   "Carrier_49_Slot2_Input" AT %IW2814 : Word;   // SLOT 2 INPUT WORD
   "Carrier_49_CrashDetectSW" AT %I2814.0 : Bool;   // CRASH DETECT SW
   "Carrier_49_SpareSafetyInput(2_1)" AT %I2814.1 : Bool;   // SPARE SAFETY INPUT
   "Carrier_49_SpareSafetyInput(2_2)" AT %I2814.2 : Bool;   // SPARE SAFETY INPUT
   "Carrier_49_SpareSafetyInput(2_3)" AT %I2814.3 : Bool;   // SPARE SAFETY INPUT
   "Carrier_49_SpareSafetyInput(2_4)" AT %I2814.4 : Bool;   // SPARE SAFETY INPUT
   "Carrier_49_SpareSafetyInput(2_5)" AT %I2814.5 : Bool;   // SPARE SAFETY INPUT
   "Carrier_49_SpareSafetyInput(2_6)" AT %I2814.6 : Bool;   // SPARE SAFETY INPUT
   "Carrier_49_SpareSafetyInput(2_7)" AT %I2814.7 : Bool;   // SPARE SAFETY INPUT
   "Carrier_49_Slot3_SafetyOutput" AT %IW2815 : Word;   // SLOT 3 SAFETY OUTPUT WORD
   "Carrier_49_Crash_Detect_OK" AT %I2815.0 : Bool;   // CARRIER CRASH DETECT
   "Carrier_49_SpareSafetyOutput(3_1)" AT %I2815.1 : Bool;   // SPARE SAFETY OUTPUT
   "Carrier_49_SpareSafetyOutput(3_2)" AT %I2815.2 : Bool;   // SPARE SAFETY OUTPUT
   "Carrier_49_SpareSafetyOutput(3_3)" AT %I2815.3 : Bool;   // SPARE SAFETY OUTPUT
   "Carrier_49_SpareSafetyOutput(3_4)" AT %I2815.4 : Bool;   // SPARE SAFETY OUTPUT
   "Carrier_49_SpareSafetyOutput(3_5)" AT %I2815.5 : Bool;   // SPARE SAFETY OUTPUT
   "Carrier_49_SpareSafetyOutput(3_6)" AT %I2815.6 : Bool;   // SPARE SAFETY OUTPUT
   "Carrier_49_SpareSafetyOutput(3_7)" AT %I2815.7 : Bool;   // SPARE SAFETY OUTPUT
   "Carrier_49_Slot4_Input" AT %IW2816 : Word;   // SLOT 4 INPUT WORD
   "Carrier_49_480VPowerOn_MDCB1" AT %I2816.0 : Bool;   // 480 VAC POWER ON MDCB 1
   "Carrier_49_SpareInput(4_1)" AT %I2816.1 : Bool;   // SPARE INPUT
   "Carrier_49_SpareInput(4_2)" AT %I2816.2 : Bool;   // SPARE INPUT
   "Carrier_49_SitopSelectStatus" AT %I2816.3 : Bool;   // SITOP SELECT STATUS
   "Carrier_49_DCsupplyOnPSCB2" AT %I2816.4 : Bool;   // DC SUPPLY ON PSCB 2
   "Carrier_49_SpareInput(4_5)" AT %I2816.5 : Bool;   // SPARE INPUT
   "Carrier_49_SpareInput(4_6)" AT %I2816.6 : Bool;   // SPARE INPUT
   "Carrier_49_SpareInput(4_7)" AT %I2816.7 : Bool;   // SPARE INPUT
   "Carrier_49_PB1_ProdHoldLH" AT %I2817.0 : Bool;   // PB 1 PRODUCTION HOLD LH
   "Carrier_49_PB2_ResetLH" AT %I2817.1 : Bool;   // PB 2 RESET LH
   "Carrier_49_PB3_ProdHoldRH" AT %I2817.2 : Bool;   // PB 3 PRODUCTION HOLD RH
   "Carrier_49_PB4_ResetRH" AT %I2817.3 : Bool;   // PB 4 RESET RH
   "Carrier_49_SpareInput(4_14)" AT %I2817.4 : Bool;   // SPARE INPUT
   "Carrier_49_SpareInput(4_15)" AT %I2817.5 : Bool;   // SPARE INPUT
   "Carrier_49_SpareInput(4_16)" AT %I2817.6 : Bool;   // SPARE INPUT
   "Carrier_49_SpareInput(4_17)" AT %I2817.7 : Bool;   // SPARE INPUT
   "Carrier_49_Slot5_Output" AT %IW2818 : Word;   // SLOT 5 OUTPUT WORD
   "Carrier_49_IRD400_HMI_24VDC_ENABLE" AT %I2818.0 : Bool;   // IRD 400 PANEL HMI 24V DC POWER
   "Carrier_49_FaultLight_LH" AT %I2818.1 : Bool;   // FAULT LIGHT LH
   "Carrier_49_RunLight_LH" AT %I2818.2 : Bool;   // RUN LIGHT LH
   "Carrier_49_FaultLight_RH" AT %I2818.3 : Bool;   // FAULT LIGHT RH
   "Carrier_49_RunLight_RH" AT %I2818.4 : Bool;   // RUN LIGHT RH
   "Carrier_49_SpareOutput(5_5)" AT %I2818.5 : Bool;   // SPARE OUTPUT
   "Carrier_49_SpareOutput(5_6)" AT %I2818.6 : Bool;   // SPARE OUTPUT
   "Carrier_49_SpareOutput(5_7)" AT %I2818.7 : Bool;   // SPARE OUTPUT
   "Carrier_49_ActualSpeed" AT %IW2820 : Word;   // ACTUAL SPEED
   "Carrier_49_CarrierDriveAlarm" AT %IW2822 : Word;   // CARRIER DRIVE ALARM
   "Carrier_49_CarrierDriveWarning" AT %IW2824 : Word;   // CARRIER DRIVE WARNING
   "Carrier_50_Status" AT %IW2850 : Word;   // CARRIER STATUS WORD
   "Carrier_50_Status.0" AT %I2850.0 : Bool;   // HEARTBEAT
   "Carrier_50_Status.1" AT %I2850.1 : Bool;   // MANUAL
   "Carrier_50_Status.2" AT %I2850.2 : Bool;   // IN_AUTO
   "Carrier_50_Status.3" AT %I2850.3 : Bool;   // POSITIONING_COMPLETE
   "Carrier_50_Status.4" AT %I2850.4 : Bool;   // PRODUCTION HOLD
   "Carrier_50_Status.5" AT %I2850.5 : Bool;   // CARRIER MOVING FORWARD
   "Carrier_50_Status.6" AT %I2850.6 : Bool;   // CARRIER MOVING REVERSE
   "Carrier_50_Status.7" AT %I2850.7 : Bool;   // CARRIER FAULT
   "Carrier_50_Status.8" AT %I2851.0 : Bool;   // CRASH DETECT TRIPPED
   "Carrier_50_Status.9" AT %I2851.1 : Bool;
   "Carrier_50_Status.10" AT %I2851.2 : Bool;
   "Carrier_50_Status.11" AT %I2851.3 : Bool;
   "Carrier_50_Status.12" AT %I2851.4 : Bool;
   "Carrier_50_Status.13" AT %I2851.5 : Bool;
   "Carrier_50_Status.14" AT %I2851.6 : Bool;
   "Carrier_50_Status.15" AT %I2851.7 : Bool;
   "Carrier_50_SDCFaultCode" AT %IW2852 : Word;   // SDC FAULT CODE
   "Carrier_50_CarrierPosition" AT %ID2854 : DWord;   // CARRIER POSITION
   "Carrier_50_CarrierNumber" AT %IW2858 : Word;   // CARRIER NUMBER
   "Carrier_50_G120DControlWord" AT %IW2860 : Word;   // G120D_STW1_CONTROL
   "Carrier_50_G120DControlWord.0" AT %I2860.0 : Bool;   // Bit_00_ON
   "Carrier_50_G120DControlWord.1" AT %I2860.1 : Bool;   // Bit_01_AUS2_INH
   "Carrier_50_G120DControlWord.2" AT %I2860.2 : Bool;   // Bit_02_AUS3_STOP
   "Carrier_50_G120DControlWord.3" AT %I2860.3 : Bool;   // Bit_03_EN
   "Carrier_50_G120DControlWord.4" AT %I2860.4 : Bool;   // Bit_04_EN_RAMP
   "Carrier_50_G120DControlWord.5" AT %I2860.5 : Bool;   // Bit_05_START_RAMP
   "Carrier_50_G120DControlWord.6" AT %I2860.6 : Bool;   // Bit_06_SETPOINT
   "Carrier_50_G120DControlWord.7" AT %I2860.7 : Bool;   // Bit_07_RESET
   "Carrier_50_G120DControlWord.8" AT %I2861.0 : Bool;   // Bit_08_JOG_R
   "Carrier_50_G120DControlWord.9" AT %I2861.1 : Bool;   // Bit_09_JOG_L
   "Carrier_50_G120DControlWord.10" AT %I2861.2 : Bool;   // Bit_10_CONTR_PLC
   "Carrier_50_G120DControlWord.11" AT %I2861.3 : Bool;   // Bit_11_REVERSE
   "Carrier_50_G120DControlWord.12" AT %I2861.4 : Bool;   // Bit_12_BRAKE_RELEASE
   "Carrier_50_G120DControlWord.13" AT %I2861.5 : Bool;   // Bit_13_DDS
   "Carrier_50_G120DControlWord.14" AT %I2861.6 : Bool;   // Bit_14_DO0
   "Carrier_50_G120DControlWord.15" AT %I2861.7 : Bool;   // Bit_15_DO1
   "Carrier_50_G120DStatusWord" AT %IW2862 : Word;   // G120D_ZSW1_STATUS
   "Carrier_50_G120DStatusWord.0" AT %I2862.0 : Bool;   // Bit_00_READY_RUN
   "Carrier_50_G120DStatusWord.1" AT %I2862.1 : Bool;   // Bit_01_READY_ON
   "Carrier_50_G120DStatusWord.2" AT %I2862.2 : Bool;   // Bit_02_ENABLE
   "Carrier_50_G120DStatusWord.3" AT %I2862.3 : Bool;   // Bit_03_FAULT
   "Carrier_50_G120DStatusWord.4" AT %I2862.4 : Bool;   // Bit_04_OFF2
   "Carrier_50_G120DStatusWord.5" AT %I2862.5 : Bool;   // Bit_05_OFF3
   "Carrier_50_G120DStatusWord.6" AT %I2862.6 : Bool;   // Bit_06_LOCK_OUT
   "Carrier_50_G120DStatusWord.7" AT %I2862.7 : Bool;   // Bit_07_WARN
   "Carrier_50_G120DStatusWord.8" AT %I2863.0 : Bool;   // Bit_08_NO_DEVIATION
   "Carrier_50_G120DStatusWord.9" AT %I2863.1 : Bool;   // Bit_09_CONTR_PLC
   "Carrier_50_G120DStatusWord.10" AT %I2863.2 : Bool;   // Bit_10_F_MAX
   "Carrier_50_G120DStatusWord.11" AT %I2863.3 : Bool;   // Bit_11_LIMIT_REACHED
   "Carrier_50_G120DStatusWord.12" AT %I2863.4 : Bool;   // Bit_12_BRAKE_OPEN
   "Carrier_50_G120DStatusWord.13" AT %I2863.5 : Bool;   // Bit_13_NO_OVERTEMP
   "Carrier_50_G120DStatusWord.14" AT %I2863.6 : Bool;   // Bit_14_CW_CCW
   "Carrier_50_G120DStatusWord.15" AT %I2863.7 : Bool;   // Bit_15_OVERL
   "Carrier_50_Slot2_Input" AT %IW2864 : Word;   // SLOT 2 INPUT WORD
   "Carrier_50_CrashDetectSW" AT %I2864.0 : Bool;   // CRASH DETECT SW
   "Carrier_50_SpareSafetyInput(2_1)" AT %I2864.1 : Bool;   // SPARE SAFETY INPUT
   "Carrier_50_SpareSafetyInput(2_2)" AT %I2864.2 : Bool;   // SPARE SAFETY INPUT
   "Carrier_50_SpareSafetyInput(2_3)" AT %I2864.3 : Bool;   // SPARE SAFETY INPUT
   "Carrier_50_SpareSafetyInput(2_4)" AT %I2864.4 : Bool;   // SPARE SAFETY INPUT
   "Carrier_50_SpareSafetyInput(2_5)" AT %I2864.5 : Bool;   // SPARE SAFETY INPUT
   "Carrier_50_SpareSafetyInput(2_6)" AT %I2864.6 : Bool;   // SPARE SAFETY INPUT
   "Carrier_50_SpareSafetyInput(2_7)" AT %I2864.7 : Bool;   // SPARE SAFETY INPUT
   "Carrier_50_Slot3_SafetyOutput" AT %IW2865 : Word;   // SLOT 3 SAFETY OUTPUT WORD
   "Carrier_50_Crash_Detect_OK" AT %I2865.0 : Bool;   // CARRIER CRASH DETECT
   "Carrier_50_SpareSafetyOutput(3_1)" AT %I2865.1 : Bool;   // SPARE SAFETY OUTPUT
   "Carrier_50_SpareSafetyOutput(3_2)" AT %I2865.2 : Bool;   // SPARE SAFETY OUTPUT
   "Carrier_50_SpareSafetyOutput(3_3)" AT %I2865.3 : Bool;   // SPARE SAFETY OUTPUT
   "Carrier_50_SpareSafetyOutput(3_4)" AT %I2865.4 : Bool;   // SPARE SAFETY OUTPUT
   "Carrier_50_SpareSafetyOutput(3_5)" AT %I2865.5 : Bool;   // SPARE SAFETY OUTPUT
   "Carrier_50_SpareSafetyOutput(3_6)" AT %I2865.6 : Bool;   // SPARE SAFETY OUTPUT
   "Carrier_50_SpareSafetyOutput(3_7)" AT %I2865.7 : Bool;   // SPARE SAFETY OUTPUT
   "Carrier_50_Slot4_Input" AT %IW2866 : Word;   // SLOT 4 INPUT WORD
   "Carrier_50_480VPowerOn_MDCB1" AT %I2866.0 : Bool;   // 480 VAC POWER ON MDCB 1
   "Carrier_50_SpareInput(4_1)" AT %I2866.1 : Bool;   // SPARE INPUT
   "Carrier_50_SpareInput(4_2)" AT %I2866.2 : Bool;   // SPARE INPUT
   "Carrier_50_SitopSelectStatus" AT %I2866.3 : Bool;   // SITOP SELECT STATUS
   "Carrier_50_DCsupplyOnPSCB2" AT %I2866.4 : Bool;   // DC SUPPLY ON PSCB 2
   "Carrier_50_SpareInput(4_5)" AT %I2866.5 : Bool;   // SPARE INPUT
   "Carrier_50_SpareInput(4_6)" AT %I2866.6 : Bool;   // SPARE INPUT
   "Carrier_50_SpareInput(4_7)" AT %I2866.7 : Bool;   // SPARE INPUT
   "Carrier_50_PB1_ProdHoldLH" AT %I2867.0 : Bool;   // PB 1 PRODUCTION HOLD LH
   "Carrier_50_PB2_ResetLH" AT %I2867.1 : Bool;   // PB 2 RESET LH
   "Carrier_50_PB3_ProdHoldRH" AT %I2867.2 : Bool;   // PB 3 PRODUCTION HOLD RH
   "Carrier_50_PB4_ResetRH" AT %I2867.3 : Bool;   // PB 4 RESET RH
   "Carrier_50_SpareInput(4_14)" AT %I2867.4 : Bool;   // SPARE INPUT
   "Carrier_50_SpareInput(4_15)" AT %I2867.5 : Bool;   // SPARE INPUT
   "Carrier_50_SpareInput(4_16)" AT %I2867.6 : Bool;   // SPARE INPUT
   "Carrier_50_SpareInput(4_17)" AT %I2867.7 : Bool;   // SPARE INPUT
   "Carrier_50_Slot5_Output" AT %IW2868 : Word;   // SLOT 5 OUTPUT WORD
   "Carrier_50_IRD400_HMI_24VDC_ENABLE" AT %I2868.0 : Bool;   // IRD 400 PANEL HMI 24V DC POWER
   "Carrier_50_FaultLight_LH" AT %I2868.1 : Bool;   // FAULT LIGHT LH
   "Carrier_50_RunLight_LH" AT %I2868.2 : Bool;   // RUN LIGHT LH
   "Carrier_50_FaultLight_RH" AT %I2868.3 : Bool;   // FAULT LIGHT RH
   "Carrier_50_RunLight_RH" AT %I2868.4 : Bool;   // RUN LIGHT RH
   "Carrier_50_SpareOutput(5_5)" AT %I2868.5 : Bool;   // SPARE OUTPUT
   "Carrier_50_SpareOutput(5_6)" AT %I2868.6 : Bool;   // SPARE OUTPUT
   "Carrier_50_SpareOutput(5_7)" AT %I2868.7 : Bool;   // SPARE OUTPUT
   "Carrier_50_ActualSpeed" AT %IW2870 : Word;   // ACTUAL SPEED
   "Carrier_50_CarrierDriveAlarm" AT %IW2872 : Word;   // CARRIER DRIVE ALARM
   "Carrier_50_CarrierDriveWarning" AT %IW2874 : Word;   // CARRIER DRIVE WARNING
   "Carrier_51_Status" AT %IW2900 : Word;   // CARRIER STATUS WORD
   "Carrier_51_Status.0" AT %I2900.0 : Bool;   // HEARTBEAT
   "Carrier_51_Status.1" AT %I2900.1 : Bool;   // MANUAL
   "Carrier_51_Status.2" AT %I2900.2 : Bool;   // IN_AUTO
   "Carrier_51_Status.3" AT %I2900.3 : Bool;   // POSITIONING_COMPLETE
   "Carrier_51_Status.4" AT %I2900.4 : Bool;   // PRODUCTION HOLD
   "Carrier_51_Status.5" AT %I2900.5 : Bool;   // CARRIER MOVING FORWARD
   "Carrier_51_Status.6" AT %I2900.6 : Bool;   // CARRIER MOVING REVERSE
   "Carrier_51_Status.7" AT %I2900.7 : Bool;   // CARRIER FAULT
   "Carrier_51_Status.8" AT %I2901.0 : Bool;   // CRASH DETECT TRIPPED
   "Carrier_51_Status.9" AT %I2901.1 : Bool;
   "Carrier_51_Status.10" AT %I2901.2 : Bool;
   "Carrier_51_Status.11" AT %I2901.3 : Bool;
   "Carrier_51_Status.12" AT %I2901.4 : Bool;
   "Carrier_51_Status.13" AT %I2901.5 : Bool;
   "Carrier_51_Status.14" AT %I2901.6 : Bool;
   "Carrier_51_Status.15" AT %I2901.7 : Bool;
   "Carrier_51_SDCFaultCode" AT %IW2902 : Word;   // SDC FAULT CODE
   "Carrier_51_CarrierPosition" AT %ID2904 : DWord;   // CARRIER POSITION
   "Carrier_51_CarrierNumber" AT %IW2908 : Word;   // CARRIER NUMBER
   "Carrier_51_G120DControlWord" AT %IW2900 : Word;   // G120D_STW1_CONTROL
   "Carrier_51_G120DControlWord.0" AT %I2900.0 : Bool;   // Bit_00_ON
   "Carrier_51_G120DControlWord.1" AT %I2900.1 : Bool;   // Bit_01_AUS2_INH
   "Carrier_51_G120DControlWord.2" AT %I2900.2 : Bool;   // Bit_02_AUS3_STOP
   "Carrier_51_G120DControlWord.3" AT %I2900.3 : Bool;   // Bit_03_EN
   "Carrier_51_G120DControlWord.4" AT %I2900.4 : Bool;   // Bit_04_EN_RAMP
   "Carrier_51_G120DControlWord.5" AT %I2900.5 : Bool;   // Bit_05_START_RAMP
   "Carrier_51_G120DControlWord.6" AT %I2900.6 : Bool;   // Bit_06_SETPOINT
   "Carrier_51_G120DControlWord.7" AT %I2900.7 : Bool;   // Bit_07_RESET
   "Carrier_51_G120DControlWord.8" AT %I2901.0 : Bool;   // Bit_08_JOG_R
   "Carrier_51_G120DControlWord.9" AT %I2901.1 : Bool;   // Bit_09_JOG_L
   "Carrier_51_G120DControlWord.10" AT %I2901.2 : Bool;   // Bit_10_CONTR_PLC
   "Carrier_51_G120DControlWord.11" AT %I2901.3 : Bool;   // Bit_11_REVERSE
   "Carrier_51_G120DControlWord.12" AT %I2901.4 : Bool;   // Bit_12_BRAKE_RELEASE
   "Carrier_51_G120DControlWord.13" AT %I2901.5 : Bool;   // Bit_13_DDS
   "Carrier_51_G120DControlWord.14" AT %I2901.6 : Bool;   // Bit_14_DO0
   "Carrier_51_G120DControlWord.15" AT %I2901.7 : Bool;   // Bit_15_DO1
   "Carrier_51_G120DStatusWord" AT %IW2902 : Word;   // G120D_ZSW1_STATUS
   "Carrier_51_G120DStatusWord.0" AT %I2902.0 : Bool;   // Bit_00_READY_RUN
   "Carrier_51_G120DStatusWord.1" AT %I2902.1 : Bool;   // Bit_01_READY_ON
   "Carrier_51_G120DStatusWord.2" AT %I2902.2 : Bool;   // Bit_02_ENABLE
   "Carrier_51_G120DStatusWord.3" AT %I2902.3 : Bool;   // Bit_03_FAULT
   "Carrier_51_G120DStatusWord.4" AT %I2902.4 : Bool;   // Bit_04_OFF2
   "Carrier_51_G120DStatusWord.5" AT %I2902.5 : Bool;   // Bit_05_OFF3
   "Carrier_51_G120DStatusWord.6" AT %I2902.6 : Bool;   // Bit_06_LOCK_OUT
   "Carrier_51_G120DStatusWord.7" AT %I2902.7 : Bool;   // Bit_07_WARN
   "Carrier_51_G120DStatusWord.8" AT %I2903.0 : Bool;   // Bit_08_NO_DEVIATION
   "Carrier_51_G120DStatusWord.9" AT %I2903.1 : Bool;   // Bit_09_CONTR_PLC
   "Carrier_51_G120DStatusWord.10" AT %I2903.2 : Bool;   // Bit_10_F_MAX
   "Carrier_51_G120DStatusWord.11" AT %I2903.3 : Bool;   // Bit_11_LIMIT_REACHED
   "Carrier_51_G120DStatusWord.12" AT %I2903.4 : Bool;   // Bit_12_BRAKE_OPEN
   "Carrier_51_G120DStatusWord.13" AT %I2903.5 : Bool;   // Bit_13_NO_OVERTEMP
   "Carrier_51_G120DStatusWord.14" AT %I2903.6 : Bool;   // Bit_14_CW_CCW
   "Carrier_51_G120DStatusWord.15" AT %I2903.7 : Bool;   // Bit_15_OVERL
   "Carrier_51_Slot2_Input" AT %IW2904 : Word;   // SLOT 2 INPUT WORD
   "Carrier_51_CrashDetectSW" AT %I2904.0 : Bool;   // CRASH DETECT SW
   "Carrier_51_SpareSafetyInput(2_1)" AT %I2904.1 : Bool;   // SPARE SAFETY INPUT
   "Carrier_51_SpareSafetyInput(2_2)" AT %I2904.2 : Bool;   // SPARE SAFETY INPUT
   "Carrier_51_SpareSafetyInput(2_3)" AT %I2904.3 : Bool;   // SPARE SAFETY INPUT
   "Carrier_51_SpareSafetyInput(2_4)" AT %I2904.4 : Bool;   // SPARE SAFETY INPUT
   "Carrier_51_SpareSafetyInput(2_5)" AT %I2904.5 : Bool;   // SPARE SAFETY INPUT
   "Carrier_51_SpareSafetyInput(2_6)" AT %I2904.6 : Bool;   // SPARE SAFETY INPUT
   "Carrier_51_SpareSafetyInput(2_7)" AT %I2904.7 : Bool;   // SPARE SAFETY INPUT
   "Carrier_51_Slot3_SafetyOutput" AT %IW2905 : Word;   // SLOT 3 SAFETY OUTPUT WORD
   "Carrier_51_Crash_Detect_OK" AT %I2905.0 : Bool;   // CARRIER CRASH DETECT
   "Carrier_51_SpareSafetyOutput(3_1)" AT %I2905.1 : Bool;   // SPARE SAFETY OUTPUT
   "Carrier_51_SpareSafetyOutput(3_2)" AT %I2905.2 : Bool;   // SPARE SAFETY OUTPUT
   "Carrier_51_SpareSafetyOutput(3_3)" AT %I2905.3 : Bool;   // SPARE SAFETY OUTPUT
   "Carrier_51_SpareSafetyOutput(3_4)" AT %I2905.4 : Bool;   // SPARE SAFETY OUTPUT
   "Carrier_51_SpareSafetyOutput(3_5)" AT %I2905.5 : Bool;   // SPARE SAFETY OUTPUT
   "Carrier_51_SpareSafetyOutput(3_6)" AT %I2905.6 : Bool;   // SPARE SAFETY OUTPUT
   "Carrier_51_SpareSafetyOutput(3_7)" AT %I2905.7 : Bool;   // SPARE SAFETY OUTPUT
   "Carrier_51_Slot4_Input" AT %IW2906 : Word;   // SLOT 4 INPUT WORD
   "Carrier_51_480VPowerOn_MDCB1" AT %I2906.0 : Bool;   // 480 VAC POWER ON MDCB 1
   "Carrier_51_SpareInput(4_1)" AT %I2906.1 : Bool;   // SPARE INPUT
   "Carrier_51_SpareInput(4_2)" AT %I2906.2 : Bool;   // SPARE INPUT
   "Carrier_51_SitopSelectStatus" AT %I2906.3 : Bool;   // SITOP SELECT STATUS
   "Carrier_51_DCsupplyOnPSCB2" AT %I2906.4 : Bool;   // DC SUPPLY ON PSCB 2
   "Carrier_51_SpareInput(4_5)" AT %I2906.5 : Bool;   // SPARE INPUT
   "Carrier_51_SpareInput(4_6)" AT %I2906.6 : Bool;   // SPARE INPUT
   "Carrier_51_SpareInput(4_7)" AT %I2906.7 : Bool;   // SPARE INPUT
   "Carrier_51_PB1_ProdHoldLH" AT %I2907.0 : Bool;   // PB 1 PRODUCTION HOLD LH
   "Carrier_51_PB2_ResetLH" AT %I2907.1 : Bool;   // PB 2 RESET LH
   "Carrier_51_PB3_ProdHoldRH" AT %I2907.2 : Bool;   // PB 3 PRODUCTION HOLD RH
   "Carrier_51_PB4_ResetRH" AT %I2907.3 : Bool;   // PB 4 RESET RH
   "Carrier_51_SpareInput(4_14)" AT %I2907.4 : Bool;   // SPARE INPUT
   "Carrier_51_SpareInput(4_15)" AT %I2907.5 : Bool;   // SPARE INPUT
   "Carrier_51_SpareInput(4_16)" AT %I2907.6 : Bool;   // SPARE INPUT
   "Carrier_51_SpareInput(4_17)" AT %I2907.7 : Bool;   // SPARE INPUT
   "Carrier_51_Slot5_Output" AT %IW2908 : Word;   // SLOT 5 OUTPUT WORD
   "Carrier_51_IRD400_HMI_24VDC_ENABLE" AT %I2908.0 : Bool;   // IRD 400 PANEL HMI 24V DC POWER
   "Carrier_51_FaultLight_LH" AT %I2908.1 : Bool;   // FAULT LIGHT LH
   "Carrier_51_RunLight_LH" AT %I2908.2 : Bool;   // RUN LIGHT LH
   "Carrier_51_FaultLight_RH" AT %I2908.3 : Bool;   // FAULT LIGHT RH
   "Carrier_51_RunLight_RH" AT %I2908.4 : Bool;   // RUN LIGHT RH
   "Carrier_51_SpareOutput(5_5)" AT %I2908.5 : Bool;   // SPARE OUTPUT
   "Carrier_51_SpareOutput(5_6)" AT %I2908.6 : Bool;   // SPARE OUTPUT
   "Carrier_51_SpareOutput(5_7)" AT %I2908.7 : Bool;   // SPARE OUTPUT
   "Carrier_51_ActualSpeed" AT %IW2920 : Word;   // ACTUAL SPEED
   "Carrier_51_CarrierDriveAlarm" AT %IW2922 : Word;   // CARRIER DRIVE ALARM
   "Carrier_51_CarrierDriveWarning" AT %IW2924 : Word;   // CARRIER DRIVE WARNING
   "Carrier_52_Status" AT %IW2950 : Word;   // CARRIER STATUS WORD
   "Carrier_52_Status.0" AT %I2950.0 : Bool;   // HEARTBEAT
   "Carrier_52_Status.1" AT %I2950.1 : Bool;   // MANUAL
   "Carrier_52_Status.2" AT %I2950.2 : Bool;   // IN_AUTO
   "Carrier_52_Status.3" AT %I2950.3 : Bool;   // POSITIONING_COMPLETE
   "Carrier_52_Status.4" AT %I2950.4 : Bool;   // PRODUCTION HOLD
   "Carrier_52_Status.5" AT %I2950.5 : Bool;   // CARRIER MOVING FORWARD
   "Carrier_52_Status.6" AT %I2950.6 : Bool;   // CARRIER MOVING REVERSE
   "Carrier_52_Status.7" AT %I2950.7 : Bool;   // CARRIER FAULT
   "Carrier_52_Status.8" AT %I2951.0 : Bool;   // CRASH DETECT TRIPPED
   "Carrier_52_Status.9" AT %I2951.1 : Bool;
   "Carrier_52_Status.10" AT %I2951.2 : Bool;
   "Carrier_52_Status.11" AT %I2951.3 : Bool;
   "Carrier_52_Status.12" AT %I2951.4 : Bool;
   "Carrier_52_Status.13" AT %I2951.5 : Bool;
   "Carrier_52_Status.14" AT %I2951.6 : Bool;
   "Carrier_52_Status.15" AT %I2951.7 : Bool;
   "Carrier_52_SDCFaultCode" AT %IW2952 : Word;   // SDC FAULT CODE
   "Carrier_52_CarrierPosition" AT %ID2954 : DWord;   // CARRIER POSITION
   "Carrier_52_CarrierNumber" AT %IW2958 : Word;   // CARRIER NUMBER
   "Carrier_52_G120DControlWord" AT %IW2960 : Word;   // G120D_STW1_CONTROL
   "Carrier_52_G120DControlWord.0" AT %I2960.0 : Bool;   // Bit_00_ON
   "Carrier_52_G120DControlWord.1" AT %I2960.1 : Bool;   // Bit_01_AUS2_INH
   "Carrier_52_G120DControlWord.2" AT %I2960.2 : Bool;   // Bit_02_AUS3_STOP
   "Carrier_52_G120DControlWord.3" AT %I2960.3 : Bool;   // Bit_03_EN
   "Carrier_52_G120DControlWord.4" AT %I2960.4 : Bool;   // Bit_04_EN_RAMP
   "Carrier_52_G120DControlWord.5" AT %I2960.5 : Bool;   // Bit_05_START_RAMP
   "Carrier_52_G120DControlWord.6" AT %I2960.6 : Bool;   // Bit_06_SETPOINT
   "Carrier_52_G120DControlWord.7" AT %I2960.7 : Bool;   // Bit_07_RESET
   "Carrier_52_G120DControlWord.8" AT %I2961.0 : Bool;   // Bit_08_JOG_R
   "Carrier_52_G120DControlWord.9" AT %I2961.1 : Bool;   // Bit_09_JOG_L
   "Carrier_52_G120DControlWord.10" AT %I2961.2 : Bool;   // Bit_10_CONTR_PLC
   "Carrier_52_G120DControlWord.11" AT %I2961.3 : Bool;   // Bit_11_REVERSE
   "Carrier_52_G120DControlWord.12" AT %I2961.4 : Bool;   // Bit_12_BRAKE_RELEASE
   "Carrier_52_G120DControlWord.13" AT %I2961.5 : Bool;   // Bit_13_DDS
   "Carrier_52_G120DControlWord.14" AT %I2961.6 : Bool;   // Bit_14_DO0
   "Carrier_52_G120DControlWord.15" AT %I2961.7 : Bool;   // Bit_15_DO1
   "Carrier_52_G120DStatusWord" AT %IW2962 : Word;   // G120D_ZSW1_STATUS
   "Carrier_52_G120DStatusWord.0" AT %I2962.0 : Bool;   // Bit_00_READY_RUN
   "Carrier_52_G120DStatusWord.1" AT %I2962.1 : Bool;   // Bit_01_READY_ON
   "Carrier_52_G120DStatusWord.2" AT %I2962.2 : Bool;   // Bit_02_ENABLE
   "Carrier_52_G120DStatusWord.3" AT %I2962.3 : Bool;   // Bit_03_FAULT
   "Carrier_52_G120DStatusWord.4" AT %I2962.4 : Bool;   // Bit_04_OFF2
   "Carrier_52_G120DStatusWord.5" AT %I2962.5 : Bool;   // Bit_05_OFF3
   "Carrier_52_G120DStatusWord.6" AT %I2962.6 : Bool;   // Bit_06_LOCK_OUT
   "Carrier_52_G120DStatusWord.7" AT %I2962.7 : Bool;   // Bit_07_WARN
   "Carrier_52_G120DStatusWord.8" AT %I2963.0 : Bool;   // Bit_08_NO_DEVIATION
   "Carrier_52_G120DStatusWord.9" AT %I2963.1 : Bool;   // Bit_09_CONTR_PLC
   "Carrier_52_G120DStatusWord.10" AT %I2963.2 : Bool;   // Bit_10_F_MAX
   "Carrier_52_G120DStatusWord.11" AT %I2963.3 : Bool;   // Bit_11_LIMIT_REACHED
   "Carrier_52_G120DStatusWord.12" AT %I2963.4 : Bool;   // Bit_12_BRAKE_OPEN
   "Carrier_52_G120DStatusWord.13" AT %I2963.5 : Bool;   // Bit_13_NO_OVERTEMP
   "Carrier_52_G120DStatusWord.14" AT %I2963.6 : Bool;   // Bit_14_CW_CCW
   "Carrier_52_G120DStatusWord.15" AT %I2963.7 : Bool;   // Bit_15_OVERL
   "Carrier_52_Slot2_Input" AT %IW2964 : Word;   // SLOT 2 INPUT WORD
   "Carrier_52_CrashDetectSW" AT %I2964.0 : Bool;   // CRASH DETECT SW
   "Carrier_52_SpareSafetyInput(2_1)" AT %I2964.1 : Bool;   // SPARE SAFETY INPUT
   "Carrier_52_SpareSafetyInput(2_2)" AT %I2964.2 : Bool;   // SPARE SAFETY INPUT
   "Carrier_52_SpareSafetyInput(2_3)" AT %I2964.3 : Bool;   // SPARE SAFETY INPUT
   "Carrier_52_SpareSafetyInput(2_4)" AT %I2964.4 : Bool;   // SPARE SAFETY INPUT
   "Carrier_52_SpareSafetyInput(2_5)" AT %I2964.5 : Bool;   // SPARE SAFETY INPUT
   "Carrier_52_SpareSafetyInput(2_6)" AT %I2964.6 : Bool;   // SPARE SAFETY INPUT
   "Carrier_52_SpareSafetyInput(2_7)" AT %I2964.7 : Bool;   // SPARE SAFETY INPUT
   "Carrier_52_Slot3_SafetyOutput" AT %IW2965 : Word;   // SLOT 3 SAFETY OUTPUT WORD
   "Carrier_52_Crash_Detect_OK" AT %I2965.0 : Bool;   // CARRIER CRASH DETECT
   "Carrier_52_SpareSafetyOutput(3_1)" AT %I2965.1 : Bool;   // SPARE SAFETY OUTPUT
   "Carrier_52_SpareSafetyOutput(3_2)" AT %I2965.2 : Bool;   // SPARE SAFETY OUTPUT
   "Carrier_52_SpareSafetyOutput(3_3)" AT %I2965.3 : Bool;   // SPARE SAFETY OUTPUT
   "Carrier_52_SpareSafetyOutput(3_4)" AT %I2965.4 : Bool;   // SPARE SAFETY OUTPUT
   "Carrier_52_SpareSafetyOutput(3_5)" AT %I2965.5 : Bool;   // SPARE SAFETY OUTPUT
   "Carrier_52_SpareSafetyOutput(3_6)" AT %I2965.6 : Bool;   // SPARE SAFETY OUTPUT
   "Carrier_52_SpareSafetyOutput(3_7)" AT %I2965.7 : Bool;   // SPARE SAFETY OUTPUT
   "Carrier_52_Slot4_Input" AT %IW2966 : Word;   // SLOT 4 INPUT WORD
   "Carrier_52_480VPowerOn_MDCB1" AT %I2966.0 : Bool;   // 480 VAC POWER ON MDCB 1
   "Carrier_52_SpareInput(4_1)" AT %I2966.1 : Bool;   // SPARE INPUT
   "Carrier_52_SpareInput(4_2)" AT %I2966.2 : Bool;   // SPARE INPUT
   "Carrier_52_SitopSelectStatus" AT %I2966.3 : Bool;   // SITOP SELECT STATUS
   "Carrier_52_DCsupplyOnPSCB2" AT %I2966.4 : Bool;   // DC SUPPLY ON PSCB 2
   "Carrier_52_SpareInput(4_5)" AT %I2966.5 : Bool;   // SPARE INPUT
   "Carrier_52_SpareInput(4_6)" AT %I2966.6 : Bool;   // SPARE INPUT
   "Carrier_52_SpareInput(4_7)" AT %I2966.7 : Bool;   // SPARE INPUT
   "Carrier_52_PB1_ProdHoldLH" AT %I2967.0 : Bool;   // PB 1 PRODUCTION HOLD LH
   "Carrier_52_PB2_ResetLH" AT %I2967.1 : Bool;   // PB 2 RESET LH
   "Carrier_52_PB3_ProdHoldRH" AT %I2967.2 : Bool;   // PB 3 PRODUCTION HOLD RH
   "Carrier_52_PB4_ResetRH" AT %I2967.3 : Bool;   // PB 4 RESET RH
   "Carrier_52_SpareInput(4_14)" AT %I2967.4 : Bool;   // SPARE INPUT
   "Carrier_52_SpareInput(4_15)" AT %I2967.5 : Bool;   // SPARE INPUT
   "Carrier_52_SpareInput(4_16)" AT %I2967.6 : Bool;   // SPARE INPUT
   "Carrier_52_SpareInput(4_17)" AT %I2967.7 : Bool;   // SPARE INPUT
   "Carrier_52_Slot5_Output" AT %IW2968 : Word;   // SLOT 5 OUTPUT WORD
   "Carrier_52_IRD400_HMI_24VDC_ENABLE" AT %I2968.0 : Bool;   // IRD 400 PANEL HMI 24V DC POWER
   "Carrier_52_FaultLight_LH" AT %I2968.1 : Bool;   // FAULT LIGHT LH
   "Carrier_52_RunLight_LH" AT %I2968.2 : Bool;   // RUN LIGHT LH
   "Carrier_52_FaultLight_RH" AT %I2968.3 : Bool;   // FAULT LIGHT RH
   "Carrier_52_RunLight_RH" AT %I2968.4 : Bool;   // RUN LIGHT RH
   "Carrier_52_SpareOutput(5_5)" AT %I2968.5 : Bool;   // SPARE OUTPUT
   "Carrier_52_SpareOutput(5_6)" AT %I2968.6 : Bool;   // SPARE OUTPUT
   "Carrier_52_SpareOutput(5_7)" AT %I2968.7 : Bool;   // SPARE OUTPUT
   "Carrier_52_ActualSpeed" AT %IW2970 : Word;   // ACTUAL SPEED
   "Carrier_52_CarrierDriveAlarm" AT %IW2972 : Word;   // CARRIER DRIVE ALARM
   "Carrier_52_CarrierDriveWarning" AT %IW2974 : Word;   // CARRIER DRIVE WARNING
   "Carrier_53_Status" AT %IW3000 : Word;   // CARRIER STATUS WORD
   "Carrier_53_Status.0" AT %I3000.0 : Bool;   // HEARTBEAT
   "Carrier_53_Status.1" AT %I3000.1 : Bool;   // MANUAL
   "Carrier_53_Status.2" AT %I3000.2 : Bool;   // IN_AUTO
   "Carrier_53_Status.3" AT %I3000.3 : Bool;   // POSITIONING_COMPLETE
   "Carrier_53_Status.4" AT %I3000.4 : Bool;   // PRODUCTION HOLD
   "Carrier_53_Status.5" AT %I3000.5 : Bool;   // CARRIER MOVING FORWARD
   "Carrier_53_Status.6" AT %I3000.6 : Bool;   // CARRIER MOVING REVERSE
   "Carrier_53_Status.7" AT %I3000.7 : Bool;   // CARRIER FAULT
   "Carrier_53_Status.8" AT %I3001.0 : Bool;   // CRASH DETECT TRIPPED
   "Carrier_53_Status.9" AT %I3001.1 : Bool;
   "Carrier_53_Status.10" AT %I3001.2 : Bool;
   "Carrier_53_Status.11" AT %I3001.3 : Bool;
   "Carrier_53_Status.12" AT %I3001.4 : Bool;
   "Carrier_53_Status.13" AT %I3001.5 : Bool;
   "Carrier_53_Status.14" AT %I3001.6 : Bool;
   "Carrier_53_Status.15" AT %I3001.7 : Bool;
   "Carrier_53_SDCFaultCode" AT %IW3002 : Word;   // SDC FAULT CODE
   "Carrier_53_CarrierPosition" AT %ID3004 : DWord;   // CARRIER POSITION
   "Carrier_53_CarrierNumber" AT %IW3008 : Word;   // CARRIER NUMBER
   "Carrier_53_G120DControlWord" AT %IW3010 : Word;   // G120D_STW1_CONTROL
   "Carrier_53_G120DControlWord.0" AT %I3010.0 : Bool;   // Bit_00_ON
   "Carrier_53_G120DControlWord.1" AT %I3010.1 : Bool;   // Bit_01_AUS2_INH
   "Carrier_53_G120DControlWord.2" AT %I3010.2 : Bool;   // Bit_02_AUS3_STOP
   "Carrier_53_G120DControlWord.3" AT %I3010.3 : Bool;   // Bit_03_EN
   "Carrier_53_G120DControlWord.4" AT %I3010.4 : Bool;   // Bit_04_EN_RAMP
   "Carrier_53_G120DControlWord.5" AT %I3010.5 : Bool;   // Bit_05_START_RAMP
   "Carrier_53_G120DControlWord.6" AT %I3010.6 : Bool;   // Bit_06_SETPOINT
   "Carrier_53_G120DControlWord.7" AT %I3010.7 : Bool;   // Bit_07_RESET
   "Carrier_53_G120DControlWord.8" AT %I3011.0 : Bool;   // Bit_08_JOG_R
   "Carrier_53_G120DControlWord.9" AT %I3011.1 : Bool;   // Bit_09_JOG_L
   "Carrier_53_G120DControlWord.10" AT %I3011.2 : Bool;   // Bit_10_CONTR_PLC
   "Carrier_53_G120DControlWord.11" AT %I3011.3 : Bool;   // Bit_11_REVERSE
   "Carrier_53_G120DControlWord.12" AT %I3011.4 : Bool;   // Bit_12_BRAKE_RELEASE
   "Carrier_53_G120DControlWord.13" AT %I3011.5 : Bool;   // Bit_13_DDS
   "Carrier_53_G120DControlWord.14" AT %I3011.6 : Bool;   // Bit_14_DO0
   "Carrier_53_G120DControlWord.15" AT %I3011.7 : Bool;   // Bit_15_DO1
   "Carrier_53_G120DStatusWord" AT %IW3012 : Word;   // G120D_ZSW1_STATUS
   "Carrier_53_G120DStatusWord.0" AT %I3012.0 : Bool;   // Bit_00_READY_RUN
   "Carrier_53_G120DStatusWord.1" AT %I3012.1 : Bool;   // Bit_01_READY_ON
   "Carrier_53_G120DStatusWord.2" AT %I3012.2 : Bool;   // Bit_02_ENABLE
   "Carrier_53_G120DStatusWord.3" AT %I3012.3 : Bool;   // Bit_03_FAULT
   "Carrier_53_G120DStatusWord.4" AT %I3012.4 : Bool;   // Bit_04_OFF2
   "Carrier_53_G120DStatusWord.5" AT %I3012.5 : Bool;   // Bit_05_OFF3
   "Carrier_53_G120DStatusWord.6" AT %I3012.6 : Bool;   // Bit_06_LOCK_OUT
   "Carrier_53_G120DStatusWord.7" AT %I3012.7 : Bool;   // Bit_07_WARN
   "Carrier_53_G120DStatusWord.8" AT %I3013.0 : Bool;   // Bit_08_NO_DEVIATION
   "Carrier_53_G120DStatusWord.9" AT %I3013.1 : Bool;   // Bit_09_CONTR_PLC
   "Carrier_53_G120DStatusWord.10" AT %I3013.2 : Bool;   // Bit_10_F_MAX
   "Carrier_53_G120DStatusWord.11" AT %I3013.3 : Bool;   // Bit_11_LIMIT_REACHED
   "Carrier_53_G120DStatusWord.12" AT %I3013.4 : Bool;   // Bit_12_BRAKE_OPEN
   "Carrier_53_G120DStatusWord.13" AT %I3013.5 : Bool;   // Bit_13_NO_OVERTEMP
   "Carrier_53_G120DStatusWord.14" AT %I3013.6 : Bool;   // Bit_14_CW_CCW
   "Carrier_53_G120DStatusWord.15" AT %I3013.7 : Bool;   // Bit_15_OVERL
   "Carrier_53_Slot2_Input" AT %IW3014 : Word;   // SLOT 2 INPUT WORD
   "Carrier_53_CrashDetectSW" AT %I3014.0 : Bool;   // CRASH DETECT SW
   "Carrier_53_SpareSafetyInput(2_1)" AT %I3014.1 : Bool;   // SPARE SAFETY INPUT
   "Carrier_53_SpareSafetyInput(2_2)" AT %I3014.2 : Bool;   // SPARE SAFETY INPUT
   "Carrier_53_SpareSafetyInput(2_3)" AT %I3014.3 : Bool;   // SPARE SAFETY INPUT
   "Carrier_53_SpareSafetyInput(2_4)" AT %I3014.4 : Bool;   // SPARE SAFETY INPUT
   "Carrier_53_SpareSafetyInput(2_5)" AT %I3014.5 : Bool;   // SPARE SAFETY INPUT
   "Carrier_53_SpareSafetyInput(2_6)" AT %I3014.6 : Bool;   // SPARE SAFETY INPUT
   "Carrier_53_SpareSafetyInput(2_7)" AT %I3014.7 : Bool;   // SPARE SAFETY INPUT
   "Carrier_53_Slot3_SafetyOutput" AT %IW3015 : Word;   // SLOT 3 SAFETY OUTPUT WORD
   "Carrier_53_Crash_Detect_OK" AT %I3015.0 : Bool;   // CARRIER CRASH DETECT
   "Carrier_53_SpareSafetyOutput(3_1)" AT %I3015.1 : Bool;   // SPARE SAFETY OUTPUT
   "Carrier_53_SpareSafetyOutput(3_2)" AT %I3015.2 : Bool;   // SPARE SAFETY OUTPUT
   "Carrier_53_SpareSafetyOutput(3_3)" AT %I3015.3 : Bool;   // SPARE SAFETY OUTPUT
   "Carrier_53_SpareSafetyOutput(3_4)" AT %I3015.4 : Bool;   // SPARE SAFETY OUTPUT
   "Carrier_53_SpareSafetyOutput(3_5)" AT %I3015.5 : Bool;   // SPARE SAFETY OUTPUT
   "Carrier_53_SpareSafetyOutput(3_6)" AT %I3015.6 : Bool;   // SPARE SAFETY OUTPUT
   "Carrier_53_SpareSafetyOutput(3_7)" AT %I3015.7 : Bool;   // SPARE SAFETY OUTPUT
   "Carrier_53_Slot4_Input" AT %IW3016 : Word;   // SLOT 4 INPUT WORD
   "Carrier_53_480VPowerOn_MDCB1" AT %I3016.0 : Bool;   // 480 VAC POWER ON MDCB 1
   "Carrier_53_SpareInput(4_1)" AT %I3016.1 : Bool;   // SPARE INPUT
   "Carrier_53_SpareInput(4_2)" AT %I3016.2 : Bool;   // SPARE INPUT
   "Carrier_53_SitopSelectStatus" AT %I3016.3 : Bool;   // SITOP SELECT STATUS
   "Carrier_53_DCsupplyOnPSCB2" AT %I3016.4 : Bool;   // DC SUPPLY ON PSCB 2
   "Carrier_53_SpareInput(4_5)" AT %I3016.5 : Bool;   // SPARE INPUT
   "Carrier_53_SpareInput(4_6)" AT %I3016.6 : Bool;   // SPARE INPUT
   "Carrier_53_SpareInput(4_7)" AT %I3016.7 : Bool;   // SPARE INPUT
   "Carrier_53_PB1_ProdHoldLH" AT %I3017.0 : Bool;   // PB 1 PRODUCTION HOLD LH
   "Carrier_53_PB2_ResetLH" AT %I3017.1 : Bool;   // PB 2 RESET LH
   "Carrier_53_PB3_ProdHoldRH" AT %I3017.2 : Bool;   // PB 3 PRODUCTION HOLD RH
   "Carrier_53_PB4_ResetRH" AT %I3017.3 : Bool;   // PB 4 RESET RH
   "Carrier_53_SpareInput(4_14)" AT %I3017.4 : Bool;   // SPARE INPUT
   "Carrier_53_SpareInput(4_15)" AT %I3017.5 : Bool;   // SPARE INPUT
   "Carrier_53_SpareInput(4_16)" AT %I3017.6 : Bool;   // SPARE INPUT
   "Carrier_53_SpareInput(4_17)" AT %I3017.7 : Bool;   // SPARE INPUT
   "Carrier_53_Slot5_Output" AT %IW3018 : Word;   // SLOT 5 OUTPUT WORD
   "Carrier_53_IRD400_HMI_24VDC_ENABLE" AT %I3018.0 : Bool;   // IRD 400 PANEL HMI 24V DC POWER
   "Carrier_53_FaultLight_LH" AT %I3018.1 : Bool;   // FAULT LIGHT LH
   "Carrier_53_RunLight_LH" AT %I3018.2 : Bool;   // RUN LIGHT LH
   "Carrier_53_FaultLight_RH" AT %I3018.3 : Bool;   // FAULT LIGHT RH
   "Carrier_53_RunLight_RH" AT %I3018.4 : Bool;   // RUN LIGHT RH
   "Carrier_53_SpareOutput(5_5)" AT %I3018.5 : Bool;   // SPARE OUTPUT
   "Carrier_53_SpareOutput(5_6)" AT %I3018.6 : Bool;   // SPARE OUTPUT
   "Carrier_53_SpareOutput(5_7)" AT %I3018.7 : Bool;   // SPARE OUTPUT
   "Carrier_53_ActualSpeed" AT %IW3020 : Word;   // ACTUAL SPEED
   "Carrier_53_CarrierDriveAlarm" AT %IW3022 : Word;   // CARRIER DRIVE ALARM
   "Carrier_53_CarrierDriveWarning" AT %IW3024 : Word;   // CARRIER DRIVE WARNING
   "Carrier_54_Status" AT %IW3050 : Word;   // CARRIER STATUS WORD
   "Carrier_54_Status.0" AT %I3050.0 : Bool;   // HEARTBEAT
   "Carrier_54_Status.1" AT %I3050.1 : Bool;   // MANUAL
   "Carrier_54_Status.2" AT %I3050.2 : Bool;   // IN_AUTO
   "Carrier_54_Status.3" AT %I3050.3 : Bool;   // POSITIONING_COMPLETE
   "Carrier_54_Status.4" AT %I3050.4 : Bool;   // PRODUCTION HOLD
   "Carrier_54_Status.5" AT %I3050.5 : Bool;   // CARRIER MOVING FORWARD
